(* CODESYS project Revisora.project (continued)

// NETWORK 17
//   TD_injecaoAr.Q: gets TRUE delay time after a rising edge at IN
_ft2(CLK := principal.IP);
_w3 := TD_injecaoAr.Q OR _ft2.Q;
injecaoAr.IP R= _w3;
injecaoTpoOff R= _w3;

// NETWORK 18
// // Desliga o ar pelo tempo
//   tpoArAtivo: =================== Alterações ===================
TD_arAtivo(IN := ciclo.IP AND injecaoAr.IP, PT := tpoArAtivo); // TON

// NETWORK 19
//   TD_arAtivo.Q: gets TRUE delay time after a rising edge at IN
injecaoAr.IP R= TD_arAtivo.Q;

// NETWORK 20
//   o_injecaoAr: DQ : Regular output | AT %QX1.2
o_injecaoAr := injecaoAr.IP;

// NETWORK 21
// =============================================
// == Impressão
// =============================================
//   o_impressao: DQ : Regular output | AT %QX0.7
o_impressao := filmeMove[1].IP;

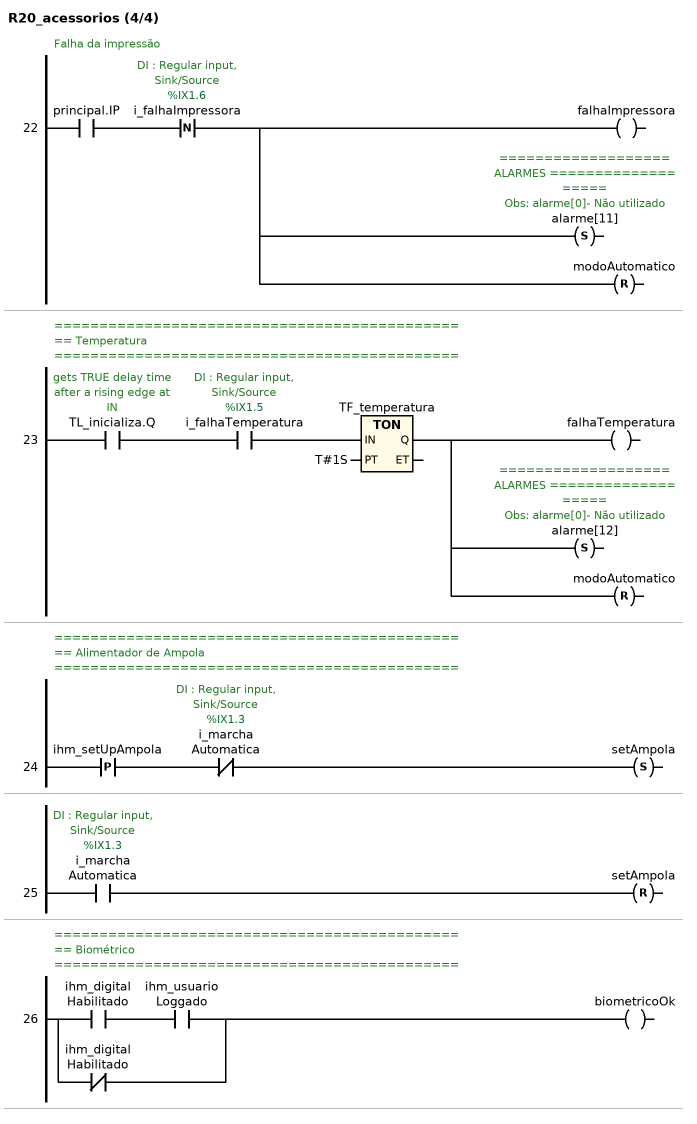
// NETWORK 22
// Falha da impressão
//   i_falhaImpressora: DI : Regular input, Sink/Source | AT %IX1.6
//   alarme[11]: =================== ALARMES =================== Obs: alarme[0]- Não utilizado
_ft3(CLK := i_falhaImpressora);
_w4 := principal.IP AND _ft3.Q;
falhaImpressora := _w4;
alarme[11] S= _w4;
modoAutomatico R= _w4;

// NETWORK 23
// =============================================
// == Temperatura
// =============================================
//   TL_inicializa.Q: gets TRUE delay time after a rising edge at IN
//   i_falhaTemperatura: DI : Regular input, Sink/Source | AT %IX1.5
//   alarme[12]: =================== ALARMES =================== Obs: alarme[0]- Não utilizado
TF_temperatura(IN := TL_inicializa.Q AND i_falhaTemperatura, PT := T#1S); // TON
falhaTemperatura := TF_temperatura.Q;
alarme[12] S= TF_temperatura.Q;
modoAutomatico R= TF_temperatura.Q;

// NETWORK 24
// =============================================
// == Alimentador de Ampola
// =============================================
//   i_marchaAutomatica: DI : Regular input, Sink/Source | AT %IX1.3
_rt3(CLK := ihm_setUpAmpola);
setAmpola S= _rt3.Q AND NOT i_marchaAutomatica;

// NETWORK 25
//   i_marchaAutomatica: DI : Regular input, Sink/Source | AT %IX1.3
setAmpola R= i_marchaAutomatica;

// NETWORK 26
// =============================================
// == Biométrico
// =============================================
biometricoOk := ihm_digitalHabilitado AND ihm_usuarioLoggado OR NOT ihm_digitalHabilitado;

END_PROGRAM

// MyController/Application/01_Machine/R06_principal
PROGRAM R06_principal
VAR
	primeiroCiclo			: BOOL;
	execMedida				: _exec_bits;
	tpoMedido				: TIME;
	T_medidaForm			: TON;
	T_inicio				: ARRAY[1..2] OF TON;
	T_selagem				: TON;
	T_arSelagem				: TON;
	T_atrasoTracao			: TON;

END_VAR
VAR // added by the converter: edge detectors and wires of the graphical bodies
    _w1, _w2, _w3, _w4, _w5, _w6, _w7, _w8, _w9, _w10, _w11, _w12, _w13 : BOOL;
    _ft1 : F_TRIG;
END_VAR

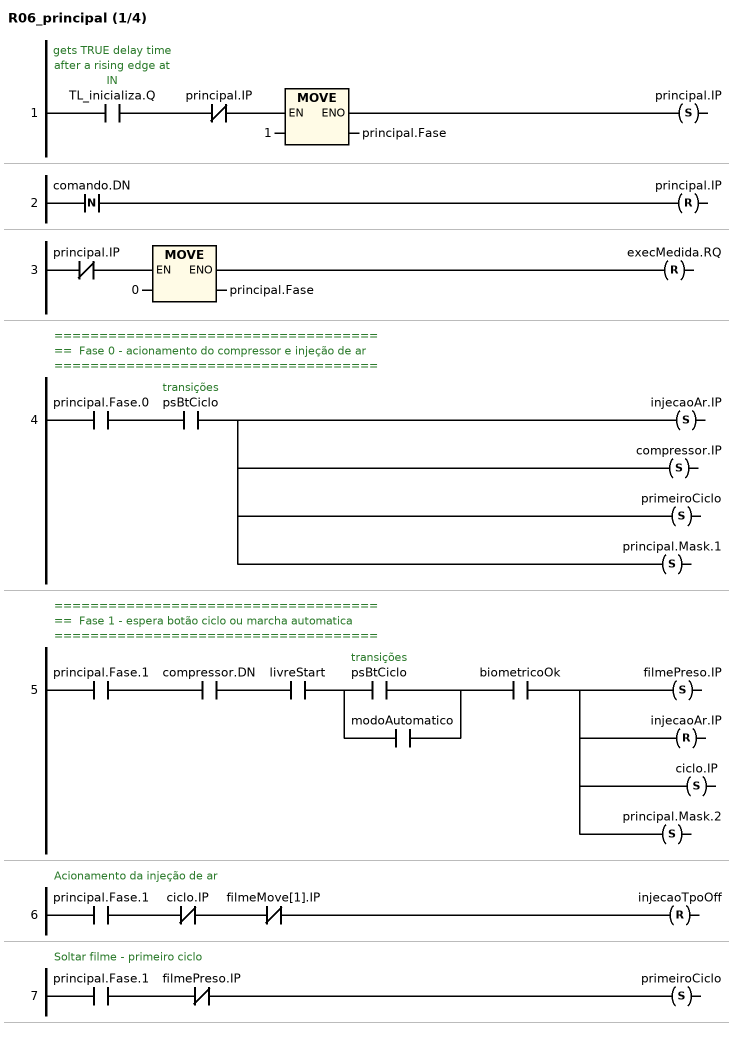
// NETWORK 1
//   TL_inicializa.Q: gets TRUE delay time after a rising edge at IN
_w1 := TL_inicializa.Q AND NOT principal.IP;
IF _w1 THEN principal.Fase := 1; END_IF
principal.IP S= _w1;

// NETWORK 2
_ft1(CLK := comando.DN);
principal.IP R= _ft1.Q;

// NETWORK 3
_w2 := NOT principal.IP;
IF _w2 THEN principal.Fase := 0; END_IF
execMedida.RQ R= _w2;

// NETWORK 4
// ====================================
// ==  Fase 0 - acionamento do compressor e injeção de ar
// ====================================
//   psBtCiclo: transições
_w3 := principal.Fase.0 AND psBtCiclo;
injecaoAr.IP S= _w3;
compressor.IP S= _w3;
primeiroCiclo S= _w3;
principal.Mask.1 S= _w3;

// NETWORK 5
// ====================================
// ==  Fase 1 - espera botão ciclo ou marcha automatica
// ====================================
//   psBtCiclo: transições
_w4 := principal.Fase.1 AND compressor.DN AND livreStart AND (psBtCiclo OR modoAutomatico) AND biometricoOk;
filmePreso.IP S= _w4;
injecaoAr.IP R= _w4;
ciclo.IP S= _w4;
principal.Mask.2 S= _w4;

// NETWORK 6
// Acionamento da injeção de ar
injecaoTpoOff R= principal.Fase.1 AND NOT ciclo.IP AND NOT filmeMove[1].IP;

// NETWORK 7
// Soltar filme - primeiro ciclo
primeiroCiclo S= principal.Fase.1 AND NOT filmePreso.IP;

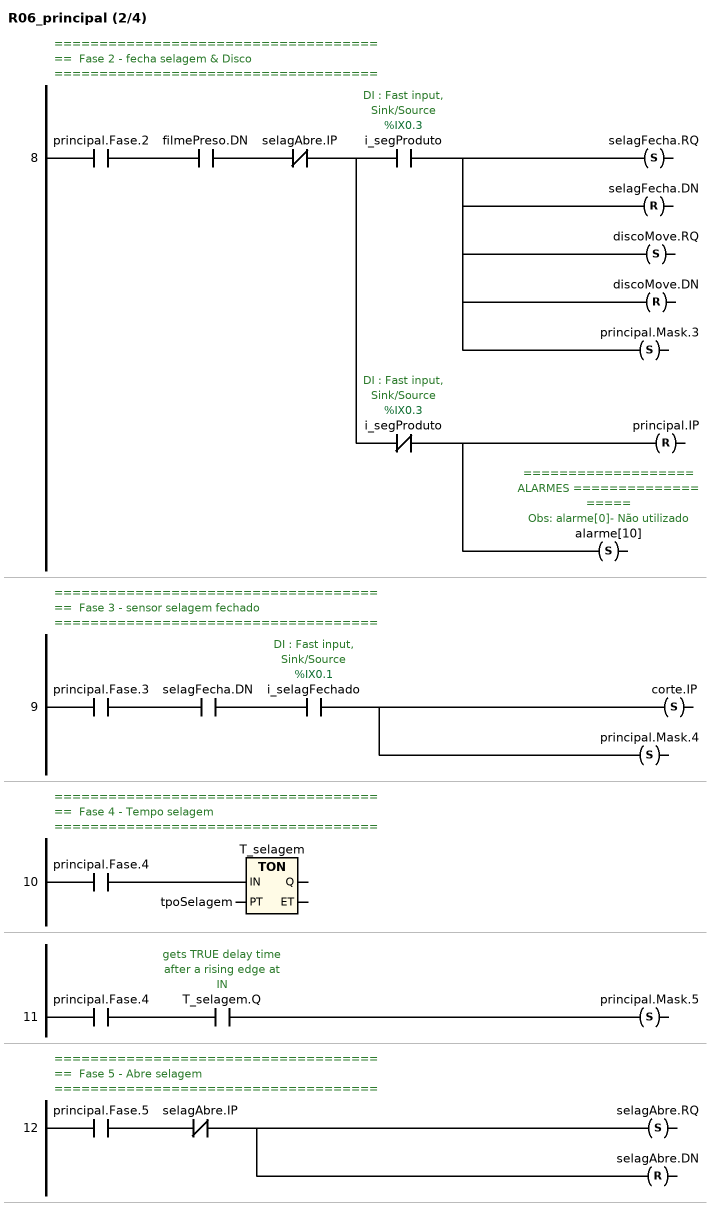
// NETWORK 8
// ====================================
// ==  Fase 2 - fecha selagem & Disco
// ====================================
//   i_segProduto: DI : Fast input, Sink/Source | AT %IX0.3
//   alarme[10]: =================== ALARMES =================== Obs: alarme[0]- Não utilizado
_w5 := principal.Fase.2 AND filmePreso.DN AND NOT selagAbre.IP;
_w6 := _w5 AND i_segProduto;
selagFecha.RQ S= _w6;
selagFecha.DN R= _w6;
discoMove.RQ S= _w6;
discoMove.DN R= _w6;
principal.Mask.3 S= _w6;
_w7 := _w5 AND NOT i_segProduto;
principal.IP R= _w7;
alarme[10] S= _w7;

// NETWORK 9
// ====================================
// ==  Fase 3 - sensor selagem fechado
// ====================================
//   i_selagFechado: DI : Fast input, Sink/Source | AT %IX0.1
_w8 := principal.Fase.3 AND selagFecha.DN AND i_selagFechado;
corte.IP S= _w8;
principal.Mask.4 S= _w8;

// NETWORK 10
// ====================================
// ==  Fase 4 - Tempo selagem
// ====================================
T_selagem(IN := principal.Fase.4, PT := tpoSelagem); // TON

// NETWORK 11
//   T_selagem.Q: gets TRUE delay time after a rising edge at IN
principal.Mask.5 S= principal.Fase.4 AND T_selagem.Q;

// NETWORK 12
// ====================================
// ==  Fase 5 - Abre selagem
// ====================================
_w9 := principal.Fase.5 AND NOT selagAbre.IP;
selagAbre.RQ S= _w9;
selagAbre.DN R= _w9;

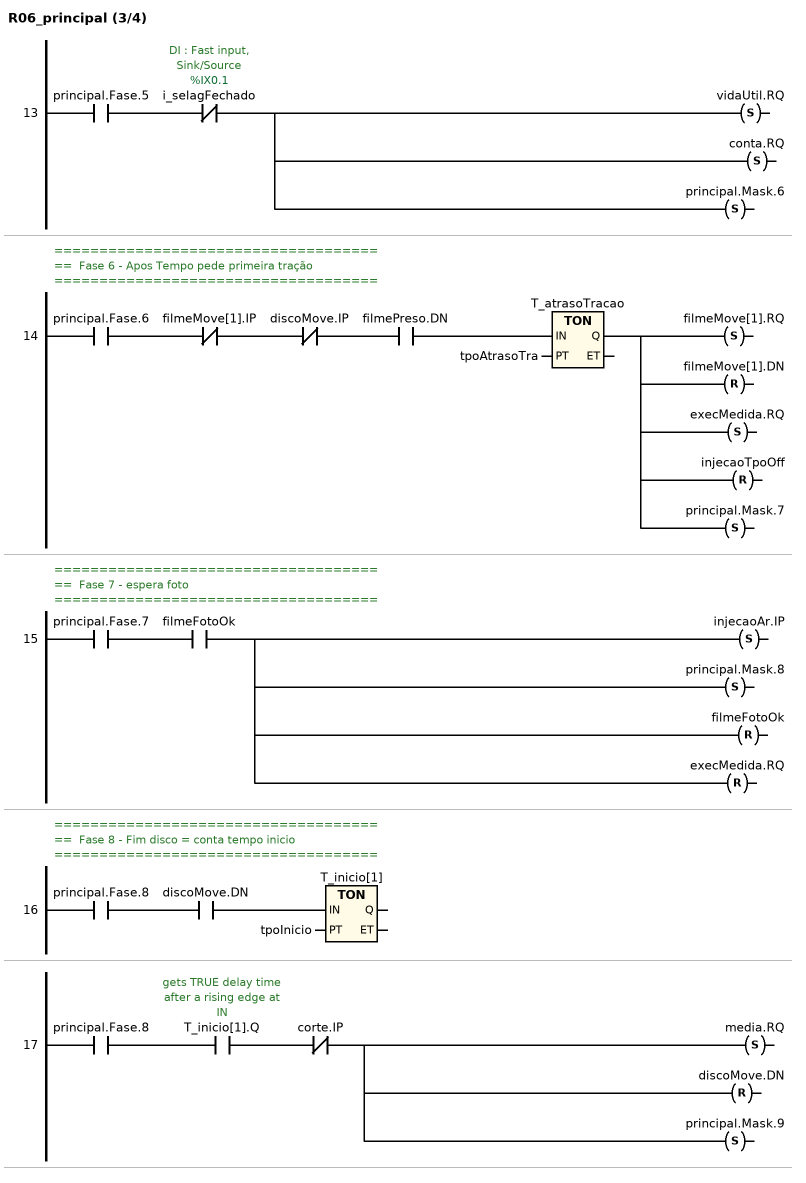
// NETWORK 13
//   i_selagFechado: DI : Fast input, Sink/Source | AT %IX0.1
_w10 := principal.Fase.5 AND NOT i_selagFechado;
vidaUtil.RQ S= _w10;
conta.RQ S= _w10;
principal.Mask.6 S= _w10;

// NETWORK 14
// ====================================
// ==  Fase 6 - Apos Tempo pede primeira tração
// ====================================
T_atrasoTracao(IN := principal.Fase.6 AND NOT filmeMove[1].IP AND NOT discoMove.IP AND filmePreso.DN, PT := tpoAtrasoTra); // TON
filmeMove[1].RQ S= T_atrasoTracao.Q;
filmeMove[1].DN R= T_atrasoTracao.Q;
execMedida.RQ S= T_atrasoTracao.Q;
injecaoTpoOff R= T_atrasoTracao.Q;
principal.Mask.7 S= T_atrasoTracao.Q;

// NETWORK 15
// ====================================
// ==  Fase 7 - espera foto
// ====================================
_w11 := principal.Fase.7 AND filmeFotoOk;
injecaoAr.IP S= _w11;
principal.Mask.8 S= _w11;
filmeFotoOk R= _w11;
execMedida.RQ R= _w11;

// NETWORK 16
// ====================================
// ==  Fase 8 - Fim disco = conta tempo inicio
// ====================================
T_inicio[1](IN := principal.Fase.8 AND discoMove.DN, PT := tpoInicio); // TON

// NETWORK 17
//   T_inicio[1].Q: gets TRUE delay time after a rising edge at IN
_w12 := principal.Fase.8 AND T_inicio[1].Q AND NOT corte.IP;
media.RQ S= _w12;
discoMove.DN R= _w12;
principal.Mask.9 S= _w12;

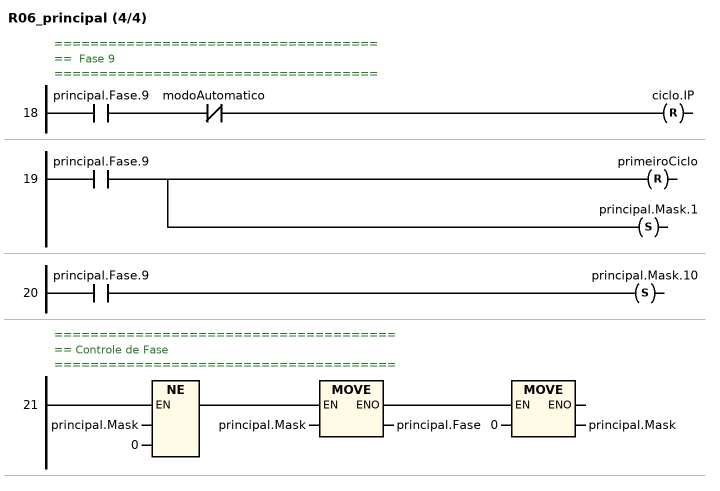
// NETWORK 18
// ====================================
// ==  Fase 9
// ====================================
ciclo.IP R= principal.Fase.9 AND NOT modoAutomatico;

// NETWORK 19
primeiroCiclo R= principal.Fase.9;
principal.Mask.1 S= principal.Fase.9;

// NETWORK 20
principal.Mask.10 S= principal.Fase.9;

// NETWORK 21
// ======================================
// == Controle de Fase
// ======================================
_w13 := principal.Mask <> 0;
IF _w13 THEN principal.Fase := principal.Mask; END_IF
IF _w13 THEN principal.Mask := 0; END_IF

END_PROGRAM

// MyController/Application/10_Relogio/AjustaDataHora
PROGRAM AjustaDataHora
VAR
	writeDateTime			: SetDateAndTime;
	readDateTime			: GetDateAndTime;
	bitScan					: BOOL;
	comOk					: BOOL;
	T_com					: TON;
END_VAR
VAR // added by the converter: edge detectors and wires of the graphical bodies
    _rt1 : R_TRIG;
END_VAR

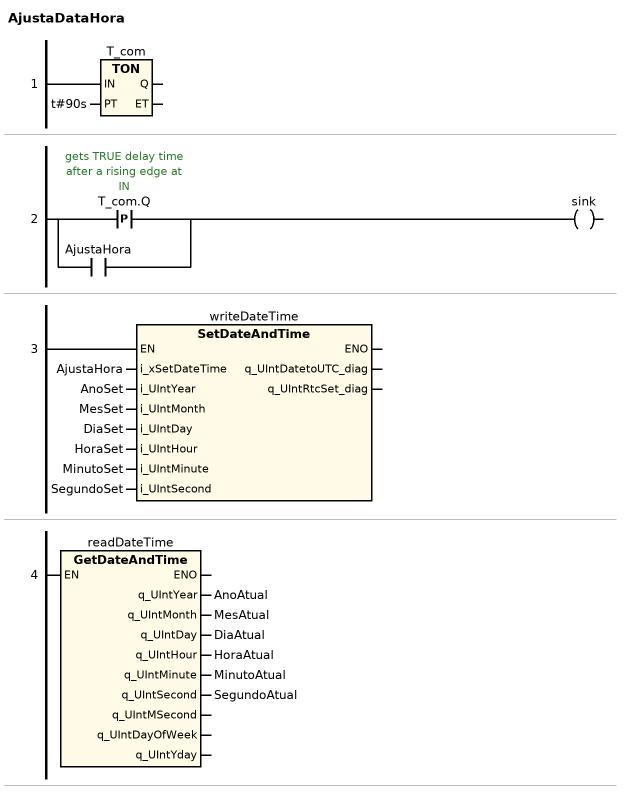
// NETWORK 1
T_com(IN := TRUE, PT := t#90s); // TON

// NETWORK 2
//   T_com.Q: gets TRUE delay time after a rising edge at IN
_rt1(CLK := T_com.Q);
sink := _rt1.Q OR AjustaHora;

// NETWORK 3
//   AnoSet: Sincroniza e ajusta o relógio da IHM
writeDateTime(
    i_xSetDateTime := AjustaHora,
    i_UIntYear := AnoSet,
    i_UIntMonth := MesSet,
    i_UIntDay := DiaSet,
    i_UIntHour := HoraSet,
    i_UIntMinute := MinutoSet,
    i_UIntSecond := SegundoSet); // SetDateAndTime

// NETWORK 4
readDateTime(
    q_UIntYear => AnoAtual,
    q_UIntMonth => MesAtual,
    q_UIntDay => DiaAtual,
    q_UIntHour => HoraAtual,
    q_UIntMinute => MinutoAtual,
    q_UIntSecond => SegundoAtual); // GetDateAndTime

END_PROGRAM

// MyController/Application/10_Relogio/SetDateAndTime
FUNCTION_BLOCK SetDateAndTime
VAR_INPUT
	i_xSetDateTime			: BOOL; (* seta novo horário na transição false para true*)
	i_UIntYear				: UINT:=2011; (*Valor para o ano a ser ajustado*)
	i_UIntMonth				: UINT:=1;(*Valor para o mes a ser ajustado*) 
	i_UIntDay				: UINT:=1;(*Valor para o dia a ser ajustado*) 
	i_UIntHour				: UINT:=0; (*Valor para a hora a ser ajustada*)
	i_UIntMinute			: UINT:=0; (*Valor para o minuto a ser ajustado*)
	i_UIntSecond			: UINT:=0;(*Valor para o segundo a ser ajustado*)
END_VAR
VAR_OUTPUT
	q_UIntDatetoUTC_diag	: UDINT; (*Status quando se =0 ok se <>0 erro nas informações de entrada*)
	q_UIntRtcSet_diag		: UDINT; (*Status quando se =0 ok se <>0 erro nas informações de entrada*)
END_VAR
VAR
	My_UTC					: DWORD; 
	MyDateTime				: SYSTIMEDATE; 
	milesec					: UINT:=0;
	dayOfWeek				: UINT:=1;
	yday					: UINT:=1;
END_VAR
VAR // added by the converter: edge detectors and wires of the graphical bodies
    _s1 : SYSTIMEDATE;
    _w1, _w2 : ANY;
END_VAR

// compose _s1 : SYSTIMEDATE
_s1.wYear := i_UIntYear;
_s1.wMonth := i_UIntMonth;
_s1.wDay := i_UIntDay;
_s1.wHour := i_UIntHour;
_s1.wMinute := i_UIntMinute;
_s1.wSecond := i_UIntSecond;
_s1.wMilliseconds := milesec;
_s1.wDayOfWeek := dayOfWeek;
_s1.wYday := yday;
MyDateTime := _s1;
_w1 := SysTimeRtcConvertDateToUtc(pDate := MyDateTime, pdwTimestampUtc := My_UTC);
q_UIntDatetoUTC_diag := _w1;
IF My_UTC <> 16#FFFFFFFF AND i_xSetDateTime THEN _w2 := SysTimeRtcSet(ulTimestamp := My_UTC); END_IF
q_UIntRtcSet_diag := _w2;
i_xSetDateTime := FALSE;

END_FUNCTION_BLOCK

// MyController/Application/10_Relogio/GetDateAndTime
FUNCTION_BLOCK GetDateAndTime
VAR_INPUT
END_VAR
VAR_OUTPUT
	q_UIntYear			: UINT; 
	q_UIntMonth			: UINT; 
	q_UIntDay			: UINT; 
	q_UIntHour			: UINT; 
	q_UIntMinute		: UINT; 
	q_UIntSecond		: UINT; 
	q_UIntMSecond		: UINT; 
	q_UIntDayOfWeek		: UINT; 
	q_UIntYday			: UINT;
END_VAR
VAR
	Ctrl_DateTime		: SYSTIMEDATE; 
	// SysTimeRtcGet operation diag 
	GetTimeResult		: UDINT; 
// SysTimeRtcConvertUtcToDate operation diag 
	UTCtoDate_diag		: UDINT; 
END_VAR
VAR // added by the converter: edge detectors and wires of the graphical bodies
    _w1, _w2 : ANY;
END_VAR

_w1 := SysTimeRtcGet(pResult := GetTimeResult);
_w2 := SysTimeRtcConvertUtcToDate(dwTimestampUtc := _w1, pDate := Ctrl_DateTime);
UTCtoDate_diag := _w2;
q_UIntYear := Ctrl_DateTime.SYSTIMEDATE;
q_UIntMonth := Ctrl_DateTime.wYear;
q_UIntDay := Ctrl_DateTime.wMonth;
q_UIntHour := Ctrl_DateTime.wDay;
q_UIntMinute := Ctrl_DateTime.wHour;
q_UIntSecond := Ctrl_DateTime.wMinute;
q_UIntMSecond := Ctrl_DateTime.wSecond;
q_UIntDayOfWeek := Ctrl_DateTime.wMilliseconds;
q_UIntYday := Ctrl_DateTime.wDayOfWeek;

END_FUNCTION_BLOCK

// MyController/Application/01_Machine/R21_estatistica
PROGRAM R21_estatistica
VAR
	infoTpoEnergizado			: RTO;
	infoTpoProducao				: RTO;
	auxHrsMinEnerg				: REAL;
	auxHrsMinProd				: REAL;				
END_VAR

(*====================================
  ==  Tempo energizado
  ====================================*)
infoTpoEnergizado(IN:= TRUE,
	  			  PT:= T#60S);
				  
infoTpoEnergizado.RST:= FALSE;			  
IF infoTpoEnergizado.Q THEN
	infoTpoEnergMin:= infoTpoEnergMin + 1;
	IF infoTpoEnergMin > 59 THEN
		infoTpoEnergHrs:= infoTpoEnergHrs + 1;
		infoTpoEnergMin:= 0;
	END_IF
	
	infoTpoEnergizado.RST:= TRUE;
END_IF


(*====================================
  ==  Tempo em produção
  ====================================*)
infoTpoProducao(IN:= ciclo.IP,
	  			PT:= T#60S);
				
IF infoTpoProducao.Q THEN
	infoTpoProdMin:= infoTpoProdMin + 1;
	IF infoTpoProdMin > 59 THEN
		infoTpoProdHrs:= infoTpoProdHrs + 1;
		infoTpoProdMin:= 0;
	END_IF
	
	infoTpoProducao.RST:= TRUE;
END_IF


// Reset dos tempos
IF estatReset THEN
	infoTpoEnergHrs:= 0;
	infoTpoEnergMin:= 0;
	infoTpoProdHrs:= 0;
	infoTpoProdMin:= 0;
	infoTpoEnergizado.RST:= TRUE;
	infoTpoProducao.RST:= TRUE;
	estatReset:= FALSE;
END_IF


(*====================================
  ==  Produtividade
  ====================================*)
// Horas e minutos energizados
auxHrsMinEnerg:= 100.0 * infoTpoEnergHrs + ((100.0 * infoTpoEnergMin) / 60.0);

// Horas e minutos em produção
auxHrsMinProd:= 100.0 * infoTpoProdHrs + ((100.0 * infoTpoProdMin) / 60.0);

IF auxHrsMinEnerg = 0 THEN
	ihm_produtMedio:= 0;
ELSE
	ihm_produtMedio:= (100.0 * auxHrsMinProd) / auxHrsMinEnerg;
END_IF



(*====================================
  ==  Conta
  ====================================*)
// Conta atual e geral
IF conta.RQ THEN
	contaAtual:= contaAtual + 1;
	contaGeral:= contaGeral + 1;
	conta.RQ:= FALSE;
END_IF

// Conta atual maior que programada = gera alarme e parada
IF contaSet <> 0 THEN
	IF contaAtual >= contaSet THEN
		alarme[3]:= TRUE;
		modoAutomatico:= FALSE;
	END_IF
END_IF


// Reset contagem atual
IF contaReset THEN
	contaAtual:= 0;
	contaReset:= FALSE;
END_IF

ihm_contaAtual:= contaAtual;
ihm_contaGeral:= contaGeral;

END_PROGRAM

// MyController/Application/11_FB/RTO
FUNCTION_BLOCK RTO
VAR_INPUT
	IN				: BOOL;
	PT				: TIME;
	RST				: BOOL;
END_VAR
VAR_OUTPUT
	Q				: BOOL;
	ACC				: TIME;
END_VAR
VAR
	auxIn			: BOOL;
	auxAcc			: TIME;
	timer			: TON;
END_VAR

IF IN AND NOT Q THEN
    ACC:= auxAcc + timer.ET;
    auxIn:= true;
end_if;

if not IN then
    auxAcc:= ACC;
    auxIn:= false;
end_if;

if ACC >= PT then
    Q:= true;
    ACC:= PT;
    auxIn:= false;
end_if;

if RST then
    Q:= false;
    ACC:= T#0s;
    auxAcc:= T#0s;
    auxIn:= false;
end_if;

timer(IN:= auxIn, PT:= T#999999S);

END_FUNCTION_BLOCK

// MyController/Application/01_Machine/R22_velocMedia
PROGRAM R22_velocMedia
VAR
	auxVelocMedia			: DINT;
	ctCiclos				: SINT;
	mediaTab				: ARRAY[0..5] OF DINT;
	mediaTpoCiclo			: DINT;
	p0						: SINT;
	T_media					: TON;
	xtr						: ARRAY[0..2] OF R_TRIG;
END_VAR

xtr[0](CLK:= compressor.DN);

IF xtr[0].Q THEN
	ctCiclos:= 0;
END_IF

media.IP:= FALSE;
IF media.RQ THEN
	mediaTpoCiclo:= TIME_TO_DINT(T_media.ET);
	media.RQ:= FALSE;
	media.IP:= TRUE;
END_IF

T_media(IN := compressor.DN AND NOT media.IP,
		PT:= T#600S);

// Carrega valores dentro da tabela		
IF media.IP THEN
	FOR p0:= 1 TO 5 DO
		mediaTab[p0 - 1]:= mediaTab[p0];
	END_FOR
	mediaTab[5]:= mediaTpoCiclo;
	
	// contagem de ciclos para efetuar a média
	IF ctCiclos < 5 THEN
		ctCiclos:= ctCiclos + 1;
	END_IF
	
	
	// Calcula média da tabela
	IF ctCiclos >= 5 THEN
		FOR p0:= 1 TO 5 DO
			IF p0 = 1 THEN
				auxVelocMedia:= 0;  // zera valor no inicio
			END_IF
			 
			auxVelocMedia:= auxVelocMedia + mediaTab[p0]; // soma todos os valores da tabela
		END_FOR
		auxVelocMedia:= auxVelocMedia / 5;
	END_IF
	
	IF auxVelocMedia <> 0 THEN
		ihm_velocMedida:= 60000 / auxVelocMedia;
	END_IF

END_IF;

END_PROGRAM

// MyController/Application/01_Machine/R98_paramFab
PROGRAM R98_paramFab
VAR
END_VAR

paramFab:= FALSE;

(*====================================
  ==  60 x 60
  ====================================*)
 Fb[0].filmeMmAposFoto:= 24;
 Fb[0].inicioAtraso:= 25;
 Fb[0].discoAtraso:= 20;
 Fb[0].inicioTracao:= 20;

 
 
(*====================================
  ==  60 x 100
  ====================================*)
 Fb[1].filmeMmAposFoto:= 24;
 Fb[1].inicioAtraso:= 25;
 Fb[1].discoAtraso:= 10;
 Fb[1].inicioTracao:= 20;
 
 
(*====================================
  ==  70 x 130
  ====================================*)
 Fb[2].filmeMmAposFoto:= 16;
 Fb[2].inicioAtraso:= 25;
 Fb[2].discoAtraso:= 0;
 Fb[2].inicioTracao:= 20;

 
 
(*====================================
  ==  X x Y
  ====================================*)
 Fb[3].filmeMmAposFoto:= 0;
 Fb[3].inicioAtraso:= 25;
 Fb[3].discoAtraso:= 0;
 Fb[3].inicioTracao:= 20;

END_PROGRAM

// MyController/Application/01_Machine/R99_calcTempos
PROGRAM R99_calcTempos
VAR
END_VAR

calcTempos:= FALSE;

// Limita os parametros de atraso de início para 10
IF Fb[numReceita].inicioAtraso < 10 THEN
	Fb[numReceita].inicioAtraso:= 10;
END_IF

IF Rc[numReceita].inicioAtraso < 10 THEN
	Rc[numReceita].inicioAtraso:= 10;
END_IF 

// Cálculo dos tempos
tpoInicio:= DINT_TO_TIME(Rc[numReceita].inicioAtraso) * 10;

tpoDisco:= DINT_TO_TIME(Rc[numReceita].discoAtraso)* 10;

tpoSelagem:= DINT_TO_TIME(M_selagTpoSelagem)* 10;

tpoAtrasoTra:= DINT_TO_TIME(Rc[numReceita].inicioTracao)* 10;

tpoInjecao:= DINT_TO_TIME(M_tpoInjecaoAr) * 10;

tpoPort:= DINT_TO_TIME(tpoAtrasPort) * 10;

tpoIniPort:= DINT_TO_TIME(inicioPort) * 10;

// Ar Ativo
tpoArAtivo:= DINT_TO_TIME(Rc[numReceita].tempoArAtivo) * 10;

END_PROGRAM

// MyController/Application/HiddenPOU
FUNCTION HiddenPOU : BOOL

VAR_INPUT
	pHiddenFunc: POINTER TO WORD;
END_VAR
VAR
	pRead: POINTER TO BYTE;
	pWrite: POINTER TO BYTE;
END_VAR

pRead := pHiddenFunc + 400;
pWrite := pHiddenFunc + 4400;
HiddenPOU := TRUE;

END_FUNCTION

// MyController/Application/Visu/Info
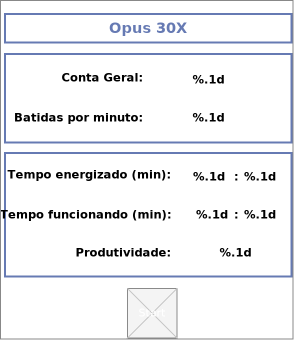
VISUALIZATION Info  // 294x340
    RoundedRectangle (4,152 288x125)
    RoundedRectangle (4,53 288x90)
    Image (127,288 50x50), "Start", image: Imagens.Botao
        OnMouseClick:  ToggleVariable=vsBtStart
    RoundedRectangle (4,13 288x30), "Opus 30X"
    Label (6,60 140x35), "Conta Geral:"
    Label (6,100 140x35), "Batidas por minuto:"
    Rectangle (151,62 115x35), "%.1d", text variable: ihm_contaGeral
    Rectangle (151,100 115x35), "%.1d", text variable: ihm_velocMedida
    Label (4,157 170x35), "Tempo energizado (min):"
    Label (4,197 170x35), "Tempo funcionando (min):"
    Rectangle (173,159 55x35), "%.1d", text variable: infoTpoEnergHrs
    Label (4,235 170x35), "Produtividade:"
    Rectangle (192,235 87x35), "%.1d", text variable: ihm_produtMedio
    Rectangle (241,159 35x35), "%.1d", text variable: infoTpoEnergMin
    Rectangle (176,197 55x35), "%.1d", text variable: infoTpoProdHrs
    Rectangle (241,197 35x35), "%.1d", text variable: infoTpoProdMin
    Label (230,159 13x35), ":"
    Label (230,197 13x35), ":"
END_VISUALIZATION

// MyController/Application/Visu/Main
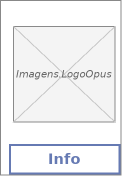
VISUALIZATION Main  // 122x176
    Image (13,26 102x96), image: Imagens.LogoOpus
    RoundedRectangle (9,144 111x30), "Info"
        OnMouseClick:  Assign=Info, Type=Assignment
END_VISUALIZATION
